(* CODESYS project Project_ROB5.project (continued)
TYPE st_CdpxButtonState :
STRUCT
	xClearError		: BOOL;
	xOperationMode	: BOOL;
	xOverview     	: BOOL;
	xUser         	: BOOL;
	xHome         	: BOOL;
	xSetupMode    	: BOOL;
	xParameter    	: BOOL;
	xSystem       	: BOOL;
	xApp_1        	: BOOL;
	xApp_2        	: BOOL;
	xStp_1        	: BOOL;
	xStp_2        	: BOOL;
	xBelt         	: BOOL;
	xApp          	: BOOL;
	xTrans_1      	: BOOL;
	xTrans_2      	: BOOL;
	xSwLanguage		: BOOL;
	xCloseDialog	: BOOL;
END_STRUCT
END_TYPE

// Data Types/SAP/ManualWork/st_MesRcvData_ManualWork
TYPE st_MesRcvData_ManualWork :
STRUCT
	stHeader		: dc_ecp.st_MES4_QueryHeader;
	sOderDes		: STRING[60];
	sPartDes		: STRING[20];
END_STRUCT
END_TYPE

// Data Types/Application/st_AppInfo
TYPE st_AppInfo :
STRUCT
	auiOperations			: ARRAY [0..15] OF UINT;
	byNumberOfOperations	: BYTE;
END_STRUCT
END_TYPE

// Data Types/SAP/sub_structures/st_Comp_Req

TYPE st_Comp_Req :
STRUCT
	sSfc	: STRING(18);
END_STRUCT
END_TYPE

// Data Types/HMI and SCADA/CDPX/st_AppSensors
TYPE st_AppSensors :
STRUCT
	xSensor		: BOOL;
	sSensor		: STRING(16);
END_STRUCT
END_TYPE

// Data Types/SAP/sub_structures/st_Comp_Res

TYPE st_Comp_Res :
STRUCT
	sOp		: STRING(4);
	sOpRev	: STRING(3);
END_STRUCT
END_TYPE

// Data Types/st_GetShuntId
TYPE st_GetShuntId :
STRUCT
	uiSourceId			: UINT;
	uiSourcePosition	: UINT;
	uiTargetId			: UINT;
	uiTargetPosition	: UINT;
END_STRUCT
END_TYPE

// Data Types/Error/st_ErrorEvent
///////////////////////////////////
///////////////////////////////////
TYPE st_ErrorEvent :
STRUCT
	/// Error ID (ID of the Errors textlist row)
	sErrorID: STRING := 'No error';
	/// Text message (It does not contains anyting, it is only to show an additional column in the visualization)
	sErrorText: STRING;
	/// String of the date and time
	sDateTime: STRING;
END_STRUCT
END_TYPE

// Data Types/HMI and SCADA/st_TransitionData
TYPE st_TransitionData :
STRUCT
	uiCondIn	: UINT;
	uiPar1		: UINT;
	uiPar2		: UINT;
	uiPar3		: UINT;
	uiPar4		: UINT;
	xAppEn		: BOOL;
	uiCondOut	: UINT;
	uiCondAbort	: UINT;
	byStopper	: BYTE;
END_STRUCT
END_TYPE

// Data Types/SAP/st_StartSfc

TYPE st_StartSfc :
STRUCT
	Req	: st_Start_Req;
	Res	: st_Start_Res;
	Com	: st_Com;
END_STRUCT
END_TYPE

// Data Types/HMI and SCADA/CDPX/st_ConveyorButtonState
TYPE st_ConveyorButtonState :
STRUCT
	xConvLeft		: BOOL;
	xConvRight		: BOOL;
	xConvSlow		: BOOL;
END_STRUCT
END_TYPE

// Global Variables/fromCDPX
{attribute 'qualified_only'}
VAR_GLOBAL
	uiMode									: UINT;
	uiDummy									: UINT;
	stCdpxButtonState						: st_CdpxButtonState;
	
	
	stHome_OperationMode_Reset		 		: st_ButtonState;
	stHome_OperationMode_Automatic		 	: st_ButtonState;
	stHome_OperationMode_Setup 				: st_ButtonState;
	stHome_OperationMode_CycleEnd 			: st_ButtonState;
	
	stSetupMode_Stopper1_Init		 		: st_ButtonState;
	stSetupMode_Stopper1_Read			 	: st_ButtonState;
	stSetupMode_Stopper1_Write 				: st_ButtonState;
	stSetupMode_Stopper1_DeleteData 		: st_ButtonState;

	stSetupMode_Stopper2_Init		 		: st_ButtonState;
	stSetupMode_Stopper2_Read			 	: st_ButtonState;
	stSetupMode_Stopper2_Write 				: st_ButtonState;
	stSetupMode_Stopper2_DeleteData 		: st_ButtonState;
	
	stInteractiveMessage_Repeat 			: st_ButtonState;
	stInteractiveMessage_Ignore	 			: st_ButtonState;
	stInteractiveMessage_Abort				: st_ButtonState;	
	stInteractiveMessage_RejectOrder		: st_ButtonState;	
	
	stManualWorkplace						: st_ManualWorkplace;
	stRobotError							: st_RobotError;	
	astStopperButton						: ARRAY [0..1] OF st_StopperButtonState;
	astAppSetting							: ARRAY [0..1] OF st_AppSettings;
	astAppButtonControl						: ARRAY [0..15] OF st_AppButtonControl;
	astTransitionTable_1					: ARRAY [0..10] OF st_TransitionData;
	astTransitionTable_2					: ARRAY [0..10] OF st_TransitionData;	
	astConveyorButtonState					: ARRAY [0..2] OF st_ConveyorButtonState; 
END_VAR

// MODULE_PLC13/Application/Variables/NVL_PLC13_SEND
VAR_GLOBAL
	Ready: BOOL := FALSE;
END_VAR

// APP_FILLING/Application/IO
//{attribute 'qualified_only'} - removed to access variables without "DigitalIO." 
VAR_GLOBAL
	// Application Type Identifier
	AppID AT %QX0.7: BOOL;
	// Push Piston forward
	PistonOn AT %QX0.1: BOOL;
	// Push Piston Backwards
	PistonOff AT %QX0.3: BOOL;
END_VAR

// Global Variables/Standards
VAR_GLOBAL
	/// First-Cycle-Flag
	xFirstCycle: BOOL := TRUE;
	/// Initialization flag
	xInit: BOOL;
	/// Station is in Initial Position
	xInitPos: BOOL;
	/// Startup like warmstart
	xSoftReset: BOOL;
	/// Application program is idle	
	xAppIdle: BOOL;
	/// Application program is busy
	xAppBusy: BOOL;
	/// Automatic Mode is active
	xAuto: BOOL;
	/// Automatic Start is enable
	xAutoEn: BOOL;
	/// Reset Mode is active
	xReset: BOOL;
	/// Reset Start is enable
	xResetEn: BOOL;
	/// Reset sequence is finished
	xResetRdy: BOOL;
	/// Manual Mode is active
	xManual: BOOL;
	/// Manual Start is enable
	xManualEn: BOOL;
	/// Teach Mode is active	
	xTeach: BOOL;
	/// Teach Start is enable
	xTeachEn: BOOL;
	/// Stop at cycle end is active	
	xCycleEnd: BOOL;
	/// Stop at cycle end is enable
	xCycleEndEn: BOOL;
	/// Reset Automatic Start flag
	xAutoReset: BOOL := FALSE;
	/// Stopper ST1 in idle state          		
	xSt1_Idle: BOOL;
	/// Stopper ST2 in idle state          		
	xSt2_Idle: BOOL;
	/// Stopper ST2 in idle state          		
	xSt3_Idle: BOOL;
	/// Resource is busy
	xBusy: BOOL;
	/// MES mode is active
	xMES: BOOL;
	/// SAP mode is active
	xSAP: BOOL;
	/// Struct with 64 Error Flags
	stError: st_Error;
	/// Structure with WinCC variables     
	stWinCC: st_WinCC;
	/// Structure with HMI variables
	stHMI: st_WinCC;
	//Semaphore for gate
	xSema : BOOL;
	// Semaphore for shunt
	xSemaShunt	: BOOL;
END_VAR

// APP_FILLING/Application/NVL_FILLING_SEND
VAR_GLOBAL
	isDone: BOOL := FALSE;
END_VAR

// MODULE_PLC13/Application/Variables/IO
VAR_GLOBAL
	

	///////////////////////////
	// Inputs
	///////////////////////////
	
	xBG20		AT %IX1.0	: BOOL;	// Stopper released
	xBG21		AT %IX1.1	: BOOL;	// Carrier available
	xBG22		AT %IX1.2	: BOOL;	// Carrier ID bit 0
	xBG23		AT %IX1.3	: BOOL;	// Carrier ID bit 1
	xBG24		AT %IX1.4	: BOOL;	// Carrier ID bit 2
	xEmg		AT %IX0.0	: BOOL;	// Emergency stop
	
	///////////////////////////
	// Outputs
	///////////////////////////	
	
	xMB20		AT %QX1.0	: BOOL;	// Release stopper
	xQA1_LEFT	AT %QX0.5	: BOOL;	// Conveyor to the left
	xQA1_RIGHT	AT %QX0.4	: BOOL;	// Conveyor to the right
	xQA1_SLOW	AT %QX0.6	: BOOL;	// Conveyor Slow
	xQA1_STOP	AT %QX0.7	: BOOL;	// Conveyor Stop
	// Application Identifier
	xAPP_ID AT %IX0.1: BOOL;
	
	
END_VAR

// Global Variables/toCDPX
{attribute 'qualified_only'}
VAR_GLOBAL
	sModule						: STRING(32);
	byOpMode					: BYTE;
	byScreenTitle				: BYTE;
	xManual						: BOOL;
	xAuto						: BOOL;
	xSAP						: BOOL;
	xMES						: BOOL;
	xDefault					: BOOL;
	auiCarrierInitNum			: ARRAY [0..1] OF UINT;
	uiNumOfApplications			: UINT;
	uiNumOfStoppers				: UINT;
	uiNumOfBelts				: UINT;
	auiCondIn					: ARRAY [0..1] OF UINT;
	auiCondOut					: ARRAY [0..1] OF UINT;
	sTime						: STRING;
	sDate						: STRING;
	stInteractiveErrors			: st_InterctiveErrors;
	astErrors					: ARRAY [1..20] OF st_Errors;
	astRfidData					: ARRAY [0..1] OF dc_ecp.st_CPF_VisuData;
	astSensorSignals			: ARRAY [0..1] OF st_StopperSensorSignals;
	astConveyorSignals			: ARRAY [0..2] OF st_ConveyorSignals;
	astAppState					: ARRAY [0..1] OF st_AppState;
	astAppControl				: ARRAY [0..1] OF st_AppControl;	
	astAppSensors				: ARRAY [0..31] OF st_AppSensors;
	auiValues					: ARRAY [0..31] OF UINT;	
	astAppControlONo: UDINT := 0;
END_VAR

// MODULE_PLC13/Application/Variables/NVL_PLC13_REC
//This gobal variable list is received via the network.
//Sender: NVL_FILLING_SEND [APP_FILLING: PLC Logic: Application]
//Protocol: UDP

VAR_GLOBAL
	isDone: BOOL := FALSE;
END_VAR

// APP_FILLING/Application/NVL_FILLING_REC
//This gobal variable list is received via the network.
//Sender: NVL_PLC13_SEND [MODULE_PLC13: PLC Logic: Application]
//Protocol: UDP

VAR_GLOBAL
	Ready: BOOL := FALSE;
END_VAR

// MODULE_PLC13/Application/Variables/NVL_PLC13_SEND
VAR_GLOBAL
	Ready: BOOL := FALSE;
END_VAR

// Global Variables/SAP
{attribute 'qualified_only'}
VAR_GLOBAL
	Start			: st_StartSfc;
	Par				: st_ParametricData;
	Comp			: st_CompleteSfc;
END_VAR

// Global Variables/SAPInit
{attribute 'qualified_only'}
VAR_GLOBAL
	Start			: st_StartSfc;
	Par				: st_ParametricData;
	Comp			: st_CompleteSfc;
END_VAR

// Global Variables/SAPHMI
{attribute 'qualified_only'}
VAR_GLOBAL
	uiOp		: UDINT;
	uiPos		: UDINT;
	sError		: STRING;
	udiSfc		: UDINT;	
END_VAR

// APP_STOPPERING/Application/IO
//{attribute 'qualified_only'} - removed to access variables without "DigitalIO." 
VAR_GLOBAL
	// Application Type Identifier
	AppID: BOOL;
	// Push Piston forward
	PistonOn: BOOL;
	// Push Piston Backwards
	PistonOff: BOOL;
	// Push second piston forwards
	Piston2On: BOOL;
	// Push second piston backwards
	Piston2Off: BOOL;
END_VAR

// APP_STOPPERING/Application/NVL_STOPPERING_SEND
VAR_GLOBAL
	isDone: BOOL := FALSE;
END_VAR

// APP_STOPPERING/Application/NVL_STOPPERING_REC
//This gobal variable list is received via the network.
//Sender: NVL_PLC13_SEND [MODULE_PLC13: PLC Logic: Application]
//Protocol: UDP

VAR_GLOBAL
	Ready: BOOL := FALSE;
END_VAR

// MODULE_PLC13/Application/Programs/MODULE_PLC13_MAIN
PROGRAM  MODULE_PLC13_MAIN
VAR
	state: UINT := 0;
	PLCid: STRING;
	RFID: dc_ecp.Dtm425;
	RfidData: dc_ecp.st_CPF_RfidData;
	ConveyorRight: BOOL;
	CarrierID: UINT;
	TIMER: TON;
	WaitTime: TIME;
	AppType: STRING;
END_VAR

CASE state OF
	
	0: // init
	IO.xMB20 := FALSE; // raise stoppper
	RFID.ClearError();
	PLCid := 'STPLC_13';
	state := 5;
	
	5: // identify
	IF IO.xAPP_ID THEN
		AppType := 'Filling';
	ELSE
		AppType := 'Stoppering';
	END_IF
		
	
	10: // wait for RFID to clear
	IF RFID.xReady THEN
		RFID.Connect(32, 0, 1);
		state:=20;
	END_IF
	
	20: // wait for RFID be ready then move conveyor
	NVL_PLC13_SEND.Ready := FALSE;
	IF RFID.xReady THEN
		IO.xMB20 := FALSE;
		IO.xQA1_RIGHT := TRUE; // Move conveyor right
		state:=30;
	END_IF
	
	30: // wait for carrier to be available
	IF IO.xBG21 THEN
		IO.xQA1_RIGHT := FALSE; // stop conveyor
		IO.xMB20 := FALSE; // lower stoppper
		state:=40;
	END_IF
	
	
	40: // wait for RFID to read then send
	NVL_PLC13_SEND.Ready := TRUE;
	IF RFID.xReady THEN
		RFID.ReadTag(uiStartAddress := 0, uiDataLength := SIZEOF(RfidData), ADR(RfidData));
		CarrierID := dc_ecp.SwapWord(RfidData.uiCarrierID); // swap bit order
		
		IF CarrierID > 0 THEN
			state:=50;
		END_IF
	END_IF
	
	
	50: // move conveyor again, give 1 sec breathing room
	IF NVL_PLC13_REC.isDone THEN
		IO.xMB20 := TRUE; // release stopper
		IF IO.xBG20 THEN // checks if stopper has been released
			IO.xQA1_RIGHT := TRUE; // move conveyor right
			WaitTime := STRING_TO_TIME('T#2000ms');
			timer(IN:=TRUE,PT:=WaitTime);
			state := 60;
		END_IF
	END_IF
	
	60: // wait for timer then restart
	IF timer.Q = TRUE THEN
		timer(IN:=FALSE);
		state := 20;
	END_IF
	
	
	
END_CASE
RFID();
timer();

END_PROGRAM

// APP_FILLING/Application/APP_FILLING_MAIN
PROGRAM APP_FILLING_MAIN
VAR
	state: UINT := 0;
	APPid: STRING;
	TIMER: TON;
	WaitTime: TIME; 
	RFID_Read : BOOL := FALSE;
END_VAR

CASE state OF
	
	0: // init
	APPid := 'APP_FILLING';
	state := 10;
	
	10: // Activate APPid & start the conveyor belt
	IO.AppID := TRUE;
	state := 15;
	
	15: // wait for module to be ready
	IF NVL_FILLING_REC.Ready THEN
		NVL_FILLING_SEND.isDone := FALSE;
		state := 20;
	END_IF
	
	20: // Push piston forward and wait 5 sec
	IO.PistonOff := FALSE;
	IO.PistonOn := TRUE;
	WaitTime := STRING_TO_TIME ('T#5000ms'); // Converts text string to time value --> WaitTime is then 5 sec
	TIMER(IN := TRUE, PT := WaitTime); // Activates the timer and the timers preset time --> The time where the piston is active
	IF Timer.Q = TRUE THEN 
		TIMER(IN := FALSE);
		state := 30;
	END_IF
	
	30: // Push piston backwards
	IO.PistonOn := FALSE;
	IO.PistonOff := TRUE;
	WaitTime := STRING_TO_TIME('T#5000ms');
	TIMER(IN := TRUE, PT := WaitTime);
	IF TIMER.Q = TRUE THEN 
		TIMER(IN := FALSE);
		state := 40;
	END_IF
	
	40: // Restart conveyor belt
	IO.PistonOff := FALSE;
	NVL_FILLING_SEND.isDone := TRUE;
	state := 15;
	
END_CASE

TIMER();

END_PROGRAM

// APP_STOPPERING/Application/APP_STOPPERING_MAIN
PROGRAM APP_STOPPERING_MAIN
VAR
	state: UINT := 0;
	APPid: STRING;
	TIMER: TON;
	WaitTime: TIME; 
	RFID_Read : BOOL := FALSE;
	TIMER2: TON := FALSE;
	TIMER3: TON := FALSE;
END_VAR

CASE state OF
	
	0: // Initilzation
	APPid := 'APP_STOPPERING';
	state := 10;
	
	10: // Activating the Stoppering application
	IO.AppID := TRUE;
	state := 15;

	15: // Checing and waiting for the module to be ready
	IF NVL_STOPPERING_REC.Ready THEN
		NVL_STOPPERING_SEND.isDone := FALSE;
		state := 20;		
	END_IF
	
	20: // Activates the first piston (in total 20 sec.) and the timer starts
	IO.PistonOn := TRUE;
	IO.PistonOff := FALSE;
	WaitTime := STRING_TO_TIME('T#20000ms');
	TIMER(IN := TRUE, PT := WaitTime);
	state := 30;
	
	30: // Checking that the first piston has been activated for 5 sec. 
	WaitTime := STRING_TO_TIME('5000ms');
	TIMER2(IN := TRUE, PT := WaitTime); 
	IF TIMER2.Q THEN // Yes - Then it activates the second piston (in total 10 sec.)
		IO.Piston2On := TRUE;
		IO.Piston2Off := FALSE;
		WaitTime := STRING_TO_TIME('T#10000');
		Timer2(IN := TRUE, PT := WaitTime);
		state := 40;
	END_IF
	
	40: // 
	IF TIMER2.Q THEN // Output variable; checking that the timer is done counting. Yes, then it deactivates second piston after 10 sec.
		IO.Piston2On := FALSE;
		IO.Piston2Off := TRUE;
		WaitTime := STRING_TO_TIME('T#5000'); // Waiting further 5 sec. + starts timer
		TIMER3(IN := TRUE, PT := WaitTime);
		state := 50;
	END_IF
	
	50: // After the last 5 sec., the first piston deactivates
	IF TIMER3.Q THEN
		IO.PistonOn := FALSE;
		IO.PistonOff := TRUE;
		state := 60;
	END_IF

	60: // End the sequence
	NVL_STOPPERING_SEND.isDone := TRUE;
	IF NOT NVL_STOPPERING_REC.Ready THEN
		state := 15;
	END_IF

END_CASE

TIMER(); // For the first piston
TIMER2(); // Second piston 
TIMER3(); // Deactivating the pistons

END_PROGRAM

// Programs/Tools/ErrorFifo
FUNCTION_BLOCK ErrorFifo
VAR_INPUT
	///Input for writing into fifo
	xWrite: BOOL;
	///Input for delete from fifo
	xDelete: BOOL;
	///The error ID
	sErrorID: STRING;
END_VAR
VAR
	///Array for the error table	
	astErrorEvent: ARRAY[1..20] OF st_ErrorEvent;
	///Triger for the rising edge of writing
	rtWrite: R_TRIG;
	///Triger for the rising edge of deleting
	rtDelete: R_TRIG;
	///Variable for the FOR loop
	uiI: UINT;
	///
	dtDateTime: DATE_AND_TIME;
	///Ask the systemtime
	fbGetTime: RTCLK.GetDateAndTime;
	///Variable to store the time data
	sDate: STRING;
	sFormat: STRING;
	rtGetTime: R_TRIG;
	xWriteTrig : BOOL;
	rtGetTimeDone: R_TRIG;
END_VAR
VAR CONSTANT
	///Not used in ARRAY SIZE !!!
	cuiSize: UINT := 20;
END_VAR

//------------------------------------------------------------------------
// ErrorFifo
//------------------------------------------------------------------------


//----------------------------------------------------------------------------------------------
// Trigger for the rising edges
//----------------------------------------------------------------------------------------------
rtWrite(CLK := xWrite);
rtDelete(CLK := xDelete);

//----------------------------------------------------------------------------------------------
// Write
//----------------------------------------------------------------------------------------------

IF rtWrite.Q THEN

//Get systemtime
	fbGetTime( xExecute:= FALSE );
	
	fbGetTime(
	xExecute:= TRUE, 
	xDone=> , 
	xBusy=> , 
	xError=> , 
	eError=> , 
	dtDateAndTime=> dtDateTime , 
	eTimezone=> );

	
	
//---------------------------------------------
// Checking the tipe of the error
//---------------------------------------------		
	IF LEFT(sErrorID, 2) = 'L0' THEN		//Level 0 error
		SysMemMove(pSrc := ADR(astErrorEvent[1]), pDest := ADR(astErrorEvent[2]), udiCount := SIZEOF(astErrorEvent) - SIZEOF(st_ErrorEvent));	
		
		astErrorEvent[1].sErrorID		:= sErrorID;
		astErrorEvent[1].sDateTime		:= sDate;

	ELSIF LEFT(sErrorID, 2) = 'L1' THEN		//Level 1 error
		FOR uiI := 1 TO cuiSize DO
			IF LEFT(astErrorEvent[uiI].sErrorID, 2) <> 'L0' THEN
				SysMemMove(pSrc := ADR(astErrorEvent[uiI]), pDest := ADR(astErrorEvent[uiI+1]), udiCount :=  SIZEOF(st_ErrorEvent) * (cuiSize-uiI-1));
		
				astErrorEvent[uiI].sErrorID		:= sErrorID;
				astErrorEvent[uiI].sDateTime	:= sDate;
				EXIT;
			END_IF
		END_FOR

	ELSIF LEFT(sErrorID, 2) = 'L2' THEN		//Level 2 error
		FOR uiI := 1 TO cuiSize DO
			IF LEFT(astErrorEvent[uiI].sErrorID, 2) <> 'L0' AND LEFT(astErrorEvent[uiI].sErrorID, 2) <> 'L1' THEN
				SysMemMove(pSrc := ADR(astErrorEvent[uiI]), pDest := ADR(astErrorEvent[uiI+1]), udiCount :=  SIZEOF(st_ErrorEvent) * (cuiSize-uiI-1));
		
				astErrorEvent[uiI].sErrorID		:= sErrorID;
				astErrorEvent[uiI].sDateTime	:= sDate;
				EXIT;
			END_IF
		END_FOR	

	END_IF
	
END_IF

sDate := DateFormat(stTime:= fbGetTime.dtDateAndTime);
//----------------------------------------------------------------------------------------------
// Delete
//----------------------------------------------------------------------------------------------
IF rtDelete.Q THEN
	FOR uiI := 1 TO cuiSize DO
		IF astErrorEvent[uiI].sErrorID = sErrorID THEN
			SysMemMove(pSrc := ADR(astErrorEvent[uiI+1]), pDest := ADR(astErrorEvent[uiI]), udiCount :=  SIZEOF(st_ErrorEvent) * (cuiSize-uiI));
			astErrorEvent[cuiSize].sErrorID		:= 'No error';
			EXIT;		
		END_IF
	END_FOR
END_IF

END_FUNCTION_BLOCK

// Programs/Tools/DateFormat
FUNCTION DateFormat : STRING
VAR_INPUT
	///Time input from ErrorFifo
	stTime: DATE_AND_TIME;
END_VAR
VAR
	///Date output in string
	sDate : STRING;
	sTemp : STRING;
	sDateTime: STRING := '';
END_VAR

//------------------------------------------------------------------------
// To show the date in the errortable in a usable format
//------------------------------------------------------------------------	

sDate := DT_TO_STRING(stTime);

//------------------------------------------------------------------------
// Cutting the days
//------------------------------------------------------------------------	

sTemp := sDate;
sDateTime := MID(STR:= sTemp, LEN:= 2, POS:= 12);
sDateTime := CONCAT(sDateTime, '/');
	
//------------------------------------------------------------------------
// Cutting the months
//------------------------------------------------------------------------		
sTemp := sDate;
sDateTime := CONCAT(sDateTime, MID(STR:= sTemp, LEN:= 2, POS:= 9));
sDateTime := CONCAT(sDateTime, '/');

//------------------------------------------------------------------------
// Cutting the years
//------------------------------------------------------------------------		

sTemp := sDate;
sDateTime := CONCAT(sDateTime, MID(STR:= sTemp, LEN:= 4, POS:= 4));
sDateTime := CONCAT(sDateTime, ' - ');	
	
//------------------------------------------------------------------------
// Cutting the hours and minutes and seconds
//------------------------------------------------------------------------	

sTemp := sDate;
sDateTime := CONCAT(sDateTime, RIGHT(STR:= sTemp, SIZE:= 8)	);

//------------------------------------------------------------------------		


	DateFormat := sDateTime;

END_FUNCTION

// Programs/Tools/MovCntr2B2M
FUNCTION_BLOCK MovCntr2B2M
VAR_INPUT
	/// Flag to Reset Error
	xQuit: BOOL;
	/// Enable error reset flag
	xQuitEN: BOOL;
	/// Enable error control
	xEnable: BOOL;
	/// Limit switch for movement 1 (M1 <--> B1) 
	xB1: BOOL;
	/// Limit switch for movement 2 (M2 <--> B2) 
	xB2: BOOL;
	/// Actor Signal for movement 1 (M1 <--> B1) 
	xM1: BOOL;
	/// Actor Signal for movement 1 (M2 <--> B2) 
	xM2: BOOL;
	/// Timeout-Time for movement 1	
	T1: TIME;
	/// Timeout-Time for movement 2
	T2: TIME;
END_VAR
VAR
	/// Timeout timer for movement 1
	TON1: TON;
	/// Timeout timer for movement 2
	TON2: TON;
	/// SR FlipFlop for Err1
	RS1: RS;
	/// SR FlipFlop for Err2
	RS2: RS;
END_VAR
VAR_OUTPUT
	/// Timeout movement 1
	xErr1: BOOL;
	/// Timeout movement 2 
	xErr2: BOOL;
END_VAR

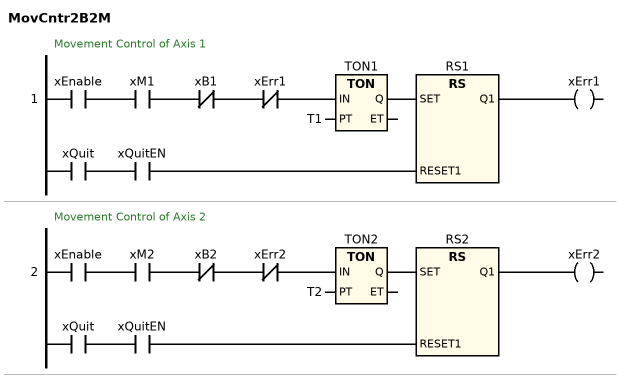
// NETWORK 1
// Movement Control of Axis 1
TON1(IN := xEnable AND xM1 AND NOT xB1 AND NOT xErr1, PT := T1); // TON
RS1(SET := TON1.Q, RESET1 := xQuit AND xQuitEN); // RS
xErr1 := RS1.Q1;

// NETWORK 2
// Movement Control of Axis 2
TON2(IN := xEnable AND xM2 AND NOT xB2 AND NOT xErr2, PT := T2); // TON
RS2(SET := TON2.Q, RESET1 := xQuit AND xQuitEN); // RS
xErr2 := RS2.Q1;

END_FUNCTION_BLOCK

// Programs/Visu/VisuProgramStp
PROGRAM  VisuProgramStp
VAR
	blBlink	: BLINK;
	t: TIME;
	uiNumOfApplications	: UINT:= 1;
	uiNumOfStoppers		: UINT:= 1;
	rtConvR				: R_TRIG;
	rtConvL				: R_TRIG;
	rtConvS				: R_TRIG;
	byActiveMainScreen	: BYTE;
	byActiveSubScreen	: BYTE;
	byScreenTitle		: BYTE;
	uiI					: UINT;
	astErrorEvents		: ARRAY [1..20] OF st_ErrorEvent;
	rtTime				: R_TRIG;
	fbGetTime: RTCLK.GetDateAndTime;
	sDate: STRING;
	dtTime	: DATE_AND_TIME;
	uiCarrierInitNum: UINT;
	xCarrierInit: BOOL;
	tonDefErr: TON;
	tonMesErr: TON;
	tonSapErr: TON;
	
	stRfidCdpx	: dc_ecp.st_CPF_RfidData;
	astAppControlONo: UDINT;
END_VAR

byActiveMainScreen	:= BOOL_TO_BYTE(fromCDPX.stCdpxButtonState.xHome)*0 + BOOL_TO_BYTE(fromCDPX.stCdpxButtonState.xSetupMode)*1 + BOOL_TO_BYTE(fromCDPX.stCdpxButtonState.xParameter)*2 + BOOL_TO_BYTE(fromCDPX.stCdpxButtonState.xSystem)*3;
byActiveSubScreen	:= BOOL_TO_BYTE(fromCDPX.stCdpxButtonState.xOperationMode)*0 + BOOL_TO_BYTE(fromCDPX.stCdpxButtonState.xApp_1)*0 +  BOOL_TO_BYTE(fromCDPX.stCdpxButtonState.xApp)*0 + BOOL_TO_BYTE(fromCDPX.stCdpxButtonState.xSystem)*0 + BOOL_TO_BYTE(fromCDPX.stCdpxButtonState.xOverview)*1 + BOOL_TO_BYTE(fromCDPX.stCdpxButtonState.xApp_2)*1 +  BOOL_TO_BYTE(fromCDPX.stCdpxButtonState.xTrans_1)*1 + BOOL_TO_BYTE(fromCDPX.stCdpxButtonState.xUser)*2 + BOOL_TO_BYTE(fromCDPX.stCdpxButtonState.xBelt)*2 +  BOOL_TO_BYTE(fromCDPX.stCdpxButtonState.xTrans_2)*2 + BOOL_TO_BYTE(fromCDPX.stCdpxButtonState.xStp_1)*3+ BOOL_TO_BYTE(fromCDPX.stCdpxButtonState.xStp_2)*4;
byScreenTitle 		:= byActiveMainScreen* 10 + byActiveSubScreen  ;

dtTime := fbGetTime.dtDateAndTime;
rtTime(CLK:= fbGetTime.xDone);
IF rtTime.Q THEN
sDate := DateFormat(stTime:= dtTime);
END_IF
fbGetTime( xExecute:= NOT fbGetTime.xDone);
fbGetTime( xExecute:= fbGetTime.xDone);

//////////////////////////////////
//			from CDPX			//
//////////////////////////////////

IF xFirstCycle THEN
	fromCDPX.astTransitionTable_1:= astTransitionTableStopper1 ;
	fromCDPX.uiMode := 1;
ELSE	
	astTransitionTableStopper1 :=fromCDPX.astTransitionTable_1;
	Visu.byMode 			:= UINT_TO_BYTE(fromCDPX.uiMode);
END_IF

// DABO /////////////////////////////////////////////////////////////////////////
IF uiCarrierInitNum <> stpStopper1.stAppSettings.uiCarrierInitNum THEN
	uiCarrierInitNum := stpStopper1.stAppSettings.uiCarrierInitNum;
ELSIF uiCarrierInitNum <> fromCDPX.astAppSetting[0].uiCarrierInitNum THEN
	uiCarrierInitNum := fromCDPX.astAppSetting[0].uiCarrierInitNum;
END_IF

fromCDPX.astAppSetting[0].uiCarrierInitNum := uiCarrierInitNum;
SysMemCpy(pDest:= ADR(stpStopper1.stAppSettings.uiCarrierInitNum), pSrc:= ADR(uiCarrierInitNum), udiCount:= SIZEOF(uiCarrierInitNum));

IF xCarrierInit <> stpStopper1.stAppSettings.xCarrierInit THEN
	xCarrierInit := stpStopper1.stAppSettings.xCarrierInit;
ELSIF xCarrierInit <> fromCDPX.astAppSetting[0].xCarrierInit THEN
	xCarrierInit := fromCDPX.astAppSetting[0].xCarrierInit;
END_IF

fromCDPX.astAppSetting[0].xCarrierInit := xCarrierInit;
SysMemCpy(pDest:= ADR(stpStopper1.stAppSettings.xCarrierInit), pSrc:= ADR(xCarrierInit), udiCount:= SIZEOF(xCarrierInit));

SysMemCpy(pDest:= ADR(stpStopper1.stAppSettings.xActive), pSrc:= ADR(fromCDPX.astAppSetting[0].xActive), udiCount:= SIZEOF(fromCDPX.astAppSetting[0].xActive));
SysMemCpy(pDest:= ADR(stpStopper1.stAppSettings.xStopBelt), pSrc:= ADR(fromCDPX.astAppSetting[0].xStopBelt), udiCount:= SIZEOF(fromCDPX.astAppSetting[0].xStopBelt));

//////////////////////////////////////////////////////////////////////////////////
// conveyor handling
rtConvL(CLK:= fromCDPX.astConveyorButtonState[0].xConvLeft);
rtConvR(CLK:= fromCDPX.astConveyorButtonState[0].xConvRight);
rtConvS(CLK:= fromCDPX.astConveyorButtonState[0].xConvSlow);
IF rtConvL.Q THEN
	IF  stpStopper1.convConveyor.xLeft THEN
		stpStopper1.convConveyor.Stop();
	ELSE
		stpStopper1.convConveyor.RunToLeft(stpStopper1.convConveyor.xSlow);
	END_IF
END_IF
IF rtConvR.Q THEN
	IF  stpStopper1.convConveyor.xRight THEN
		stpStopper1.convConveyor.Stop();
	ELSE
		stpStopper1.convConveyor.RunToRight(stpStopper1.convConveyor.xSlow);
	END_IF
END_IF
IF rtConvS.Q THEN
	IF  stpStopper1.convConveyor.xSlow THEN
		stpStopper1.convConveyor.SpeedUp();
	ELSE
		stpStopper1.convConveyor.SlowDown();
	END_IF
END_IF

// Operation mode buttons
fromCDPX.stHome_OperationMode_Reset.xActive := xReset OR (xResetEn AND blBlink.OUT);
fromCDPX.stHome_OperationMode_Reset.xDisabled := NOT xResetEn;

fromCDPX.stHome_OperationMode_Automatic.xActive := xAuto OR (xAutoEn AND blBlink.OUT);
fromCDPX.stHome_OperationMode_Automatic.xDisabled := NOT xAutoEn AND NOT xAuto;

fromCDPX.stHome_OperationMode_Setup.xActive := xManual;
fromCDPX.stHome_OperationMode_Setup.xDisabled := NOT xManualEn AND NOT xManual;

fromCDPX.stHome_OperationMode_CycleEnd.xActive := xCycleEnd AND blBlink.OUT;
fromCDPX.stHome_OperationMode_CycleEnd.xDisabled := NOT xCycleEndEn AND NOT xCycleEnd;

stWinCC.xAuto 		:= fromCDPX.stHome_OperationMode_Automatic.xPressed;
stWinCC.xReset 		:= fromCDPX.stHome_OperationMode_Reset.xPressed;
stWinCC.xManual 	:= fromCDPX.stHome_OperationMode_Setup.xPressed;
stWinCC.xCycleEnd 	:= fromCDPX.stHome_OperationMode_CycleEnd.xPressed;
stWinCC.xQuit		:= fromCDPX.stCdpxButtonState.xClearError;

// Setup RFID buttons
fromCDPX.stSetupMode_Stopper1_Init.xActive R= stpStopper1.stpStopper.dtmRfid.xReady;
fromCDPX.stSetupMode_Stopper1_Init.xActive S= fromCDPX.stSetupMode_Stopper1_Init.xPressed;
fromCDPX.stSetupMode_Stopper1_Init.xDisabled :=  xManual;
IF fromCDPX.astStopperButton[0].xInit THEN
	stpStopper1.stpStopper.Connect(usiCanChannel := stpStopper1.usiCanChannel, usiCanNetworkId := stpStopper1.usiCanNetworkId, usiCanNodeId := stpStopper1.usiCanNodeId);
END_IF


fromCDPX.stSetupMode_Stopper1_Read.xActive R= stpStopper1.stpStopper.dtmRfid.xReady;
fromCDPX.stSetupMode_Stopper1_Read.xActive S= fromCDPX.stSetupMode_Stopper1_Read.xPressed;
fromCDPX.stSetupMode_Stopper1_Read.xDisabled := xManual;
IF fromCDPX.astStopperButton[0].xRead THEN
	stpStopper1.stpStopper.ReadRfid(pstRfidData := ADR(stRfidCdpx));
	toCDPX.astRfidData[0].uiCarrierID				:=	stRfidCdpx.uiCarrierID					 ;
	toCDPX.astRfidData[0].uiCode					:=	stRfidCdpx.uiCode						 	;
	toCDPX.astRfidData[0].uiParameter1				:=	stRfidCdpx.uiParameter1					 ;
	toCDPX.astRfidData[0].uiParameter2				:=	stRfidCdpx.uiParameter2					 ;
	toCDPX.astRfidData[0].uiParameter3				:=	stRfidCdpx.uiParameter3					 ;
	toCDPX.astRfidData[0].uiParameter4				:=	stRfidCdpx.uiParameter4					 ;
	toCDPX.astRfidData[0].stMesData.udiONo			:=	stRfidCdpx.stMesData.udiONo				 ;
	toCDPX.astRfidData[0].stMesData.udiPNo			:=	stRfidCdpx.stMesData.udiPNo				 ;
	toCDPX.astRfidData[0].stMesData.uiOpNo			:=	stRfidCdpx.stMesData.uiOpNo				 ;
	toCDPX.astRfidData[0].stMesData.uiOPos			:=	stRfidCdpx.stMesData.uiOPos				 ;
	toCDPX.astRfidData[0].stMesData.uiResourceId	:=	stRfidCdpx.stMesData.uiResourceId		 	;
	toCDPX.astRfidData[0].stSapData.sItem	 		:=	stRfidCdpx.stSapData.sItem	 			 ;
	toCDPX.astRfidData[0].stSapData.sItemRev		:=	stRfidCdpx.stSapData.sItemRev			 	;
	toCDPX.astRfidData[0].stSapData.sSfc			:=	stRfidCdpx.stSapData.sSfc				 	;
	toCDPX.astRfidData[0].stSapData.udiOp			:=	stRfidCdpx.stSapData.udiOp				 ;
	toCDPX.astRfidData[0].stSapData.udiSfc			:=	stRfidCdpx.stSapData.udiSfc				 ;
END_IF                                                	


fromCDPX.stSetupMode_Stopper1_Write.xActive R= stpStopper1.stpStopper.dtmRfid.xReady;
fromCDPX.stSetupMode_Stopper1_Write.xActive S= fromCDPX.stSetupMode_Stopper1_Write.xPressed;
fromCDPX.stSetupMode_Stopper1_Write.xDisabled := xManual;
IF fromCDPX.astStopperButton[0].xWrite THEN
	stRfidCdpx.uiCarrierID					:= toCDPX.astRfidData[0].uiCarrierID				;
	stRfidCdpx.uiCode						:= toCDPX.astRfidData[0].uiCode					;
	stRfidCdpx.uiParameter1					:= toCDPX.astRfidData[0].uiParameter1				;
	stRfidCdpx.uiParameter2					:= toCDPX.astRfidData[0].uiParameter2				;
	stRfidCdpx.uiParameter3					:= toCDPX.astRfidData[0].uiParameter3				;
	stRfidCdpx.uiParameter4					:= toCDPX.astRfidData[0].uiParameter4				;
	stRfidCdpx.stMesData.udiONo				:= toCDPX.astRfidData[0].stMesData.udiONo			;
	stRfidCdpx.stMesData.udiPNo				:= toCDPX.astRfidData[0].stMesData.udiPNo			;
	stRfidCdpx.stMesData.uiOpNo				:= toCDPX.astRfidData[0].stMesData.uiOpNo			;
	stRfidCdpx.stMesData.uiOPos				:= toCDPX.astRfidData[0].stMesData.uiOPos			;
	stRfidCdpx.stMesData.uiResourceId		:= toCDPX.astRfidData[0].stMesData.uiResourceId	;
	stRfidCdpx.stSapData.sItem	 			:= toCDPX.astRfidData[0].stSapData.sItem	 		;
	stRfidCdpx.stSapData.sItemRev			:= toCDPX.astRfidData[0].stSapData.sItemRev		;
	stRfidCdpx.stSapData.sSfc				:= toCDPX.astRfidData[0].stSapData.sSfc			;
	stRfidCdpx.stSapData.udiOp				:= toCDPX.astRfidData[0].stSapData.udiOp			;
	stRfidCdpx.stSapData.udiSfc				:= toCDPX.astRfidData[0].stSapData.udiSfc			;
	stpStopper1.stpStopper.WriteRfid(stRfidData:= stRfidCdpx);
END_IF


fromCDPX.stSetupMode_Stopper1_DeleteData.xActive := fromCDPX.stSetupMode_Stopper1_DeleteData.xPressed;
fromCDPX.stSetupMode_Stopper1_DeleteData.xDisabled := xManual;                                            
IF fromCDPX.astStopperButton[0].xDeleteData	THEN
	SysMemSet(pDest:= ADR(stpStopper1.stpStopper.stRfidVisu), udiValue:= 0, udiCount:= SIZEOF(stpStopper1.stpStopper.stRfidVisu));
	SysMemCpy(pDest:= ADR(toCDPX.astRfidData[0]), pSrc:= ADR(stpStopper1.stpStopper.stRfidVisu), udiCount:= SIZEOF(stpStopper1.stpStopper.stRfidData));	
END_IF

IF NOt xManual  THEN
	SysMemCpy(pDest:= ADR(toCDPX.astRfidData[0]), pSrc:= ADR(stpStopper1.stpStopper.stRfidVisu), udiCount:= SIZEOF(stpStopper1.stpStopper.stRfidData));	
END_IF


IF fromCDPX.astStopperButton[0].xStpMveDown	THEN
	stpStopper1.stpStopper.cpfssStopper.StayDown();
END_IF
IF fromCDPX.astStopperButton[0].xStpMveUp	THEN
	stpStopper1.stpStopper.cpfssStopper.MoveUp();
END_IF

Visu.stInteractiveError.xBtnAbort 		:= fromCDPX.stInteractiveMessage_Abort.xPressed;
Visu.stInteractiveError.xBtnIgnore 		:= fromCDPX.stInteractiveMessage_Ignore.xPressed;
Visu.stInteractiveError.xBtnRejectOrder := fromCDPX.stInteractiveMessage_RejectOrder.xPressed;
Visu.stInteractiveError.xBtnRepeat		:= fromCDPX.stInteractiveMessage_Repeat.xPressed;

blBlink(ENABLE := TRUE, TIMEHIGH := T#1S, TIMELOW := T#1S); 
	

IF Visu.byMode = 1 THEN
	xMES := TRUE;
	xSAP := FALSE;
ELSIF Visu.byMode = 2 THEN
	xMES := FALSE;
	xSAP := TRUE;
ELSE
	xMES := FALSE;
	xSAP := FALSE;
END_IF

IF NOT xAuto AND NOT xManual AND NOT xReset THEN
	Visu.byOpMode := 0;
ELSIF xReset THEN
	Visu.byOpMode := 1;
ELSIF xAuto THEN
	Visu.byOpMode := 2;
ELSIF xManual THEN
	Visu.byOpMode := 3;
END_IF


//////////////////////////////////
//			to CDPX				//
//////////////////////////////////


toCDPX.byOpMode									:= Visu.byOpMode;
toCDPX.byScreenTitle							:= byScreenTitle;
toCDPX.xManual									:= xManual;	
toCDPX.xAuto									:= xAuto;			
toCDPX.xSAP										:= xSAP;				
toCDPX.xMES										:= xMES;				
toCDPX.xDefault									:= NOT xSAP AND NOT xMES;		
toCDPX.uiNumOfApplications						:= uiNumOfApplications;				
toCDPX.uiNumOfStoppers							:= uiNumOfStoppers;						
toCDPX.sDate									:= LEFT(sDate,10);
toCDPX.sTime									:= RIGHT(sDate,8);
toCDPX.auiCondIn[0]								:= stpStopper1.uiCondIn;
toCDPX.auiCondOut[0]							:= stpStopper1.uiCondOut;


toCDPX.astSensorSignals[0].sInductive_1			:= 'xBG21';
toCDPX.astSensorSignals[0].sInductive_2			:= 'xBG22';
toCDPX.astSensorSignals[0].sInductive_3			:= 'xBG23';
toCDPX.astSensorSignals[0].sInductive_4			:= 'xBG24';
toCDPX.astSensorSignals[0].sRfid				:= 'TF80';
toCDPX.astSensorSignals[0].sStpDownOutpu		:= 'xMB20';
toCDPX.astSensorSignals[0].sStpDownSensor		:= 'xBG20';
toCDPX.astSensorSignals[0].xInductive_1			:= xBG21; 
toCDPX.astSensorSignals[0].xInductive_2			:= xBG22; 
toCDPX.astSensorSignals[0].xInductive_3			:= xBG23; 
toCDPX.astSensorSignals[0].xInductive_4			:= xBG24; 
toCDPX.astSensorSignals[0].xStpDownOutpu		:= xMB20; 
toCDPX.astSensorSignals[0].xStpDownSensor		:= xBG20;
toCDPX.astSensorSignals[0].xTagPresent			:= stpStopper1.stpStopper.dtmRfid.stState.xTagPresent;
toCDPX.astSensorSignals[0].xReady				:= stpStopper1.stpStopper.dtmRfid.xReady;
toCDPX.astSensorSignals[0].xBusy				:= NOT stpStopper1.stpStopper.dtmRfid.xReady;
toCDPX.astSensorSignals[0].xError				:= stpStopper1.stpStopper.dtmRfid.xError;
toCDPX.astSensorSignals[0].xTimeOut				:= stpStopper1.stpStopper.dtmRfid.xTimeout;
                                               
